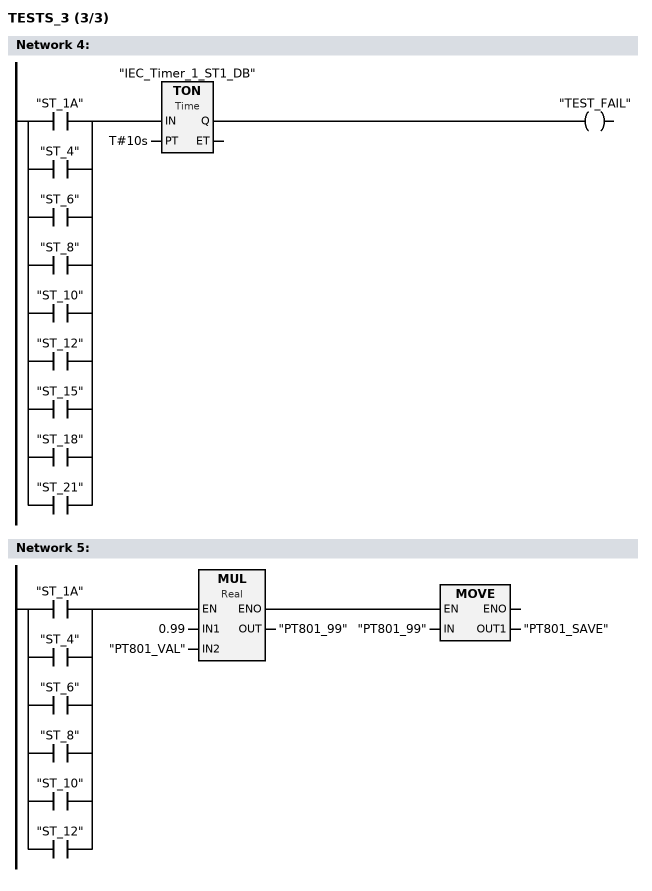
   "IEC_Timer_1_ST1_DB".TON(IN := "ST_1A" OR "ST_4" OR "ST_6" OR "ST_8" OR "ST_10" OR "ST_12" OR "ST_15" OR "ST_18" OR "ST_21",
                           PT := T#10s);
   "TEST_FAIL" := "IEC_Timer_1_ST1_DB".Q;
END_REGION

REGION Network 5
   RUNG wire#powerrail
      Contact( "ST_1A" )
      wire#w1
      { S7_Templates := "SrcType := Real" } Mul(in1 := 0.99, in2 := "PT801_VAL", out => "PT801_99")
      { S7_GenerateENO := "TRUE" } Move(in := "PT801_99", out1 => "PT801_SAVE")
   END_RUNG
   RUNG wire#powerrail
      Contact( "ST_4" )
   END_RUNG wire#w1
   RUNG wire#powerrail
      Contact( "ST_6" )
   END_RUNG wire#w1
   RUNG wire#powerrail
      Contact( "ST_8" )
   END_RUNG wire#w1
   RUNG wire#powerrail
      Contact( "ST_10" )
   END_RUNG wire#w1
   RUNG wire#powerrail
      Contact( "ST_12" )
   END_RUNG wire#w1
   // the same network as SCL:
   IF "ST_1A" OR "ST_4" OR "ST_6" OR "ST_8" OR "ST_10" OR "ST_12" THEN
       "PT801_99" := 0.99 * "PT801_VAL";
       "PT801_SAVE" := "PT801_99";
   END_IF;
END_REGION
END_FUNCTION

FUNCTION "TESTS_2" : Void   // FC18, LAD
{ S7_Optimized_Access := 'FALSE' }
VERSION : 0.1
// Test_MFC401
   VAR_TEMP   // added for the SCL form of the ladder/FBD networks
      _w1 : Bool;
      _w2 : Bool;
   END_VAR
BEGIN

REGION Network 1
   // ALARM Settings
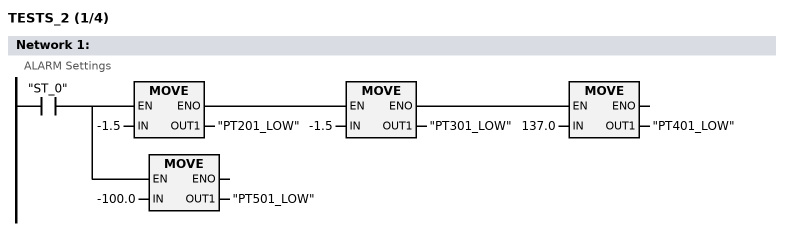
   RUNG wire#powerrail
      Contact( "ST_0" )
      wire#w1
      { S7_GenerateENO := "TRUE" } Move(in := -1.5, out1 => "PT201_LOW")
      { S7_GenerateENO := "TRUE" } Move(in := -1.5, out1 => "PT301_LOW")
      { S7_GenerateENO := "TRUE" } Move(in := 137.0, out1 => "PT401_LOW")
   END_RUNG
   RUNG wire#w1
      { S7_GenerateENO := "TRUE" } Move(in := -100.0, out1 => "PT501_LOW")
   END_RUNG
   // the same network as SCL:
   // ENO of a box is taken as its EN; it also drops when the box reports an error
   IF "ST_0" THEN
       "PT201_LOW" := -1.5;
       "PT301_LOW" := -1.5;
       "PT401_LOW" := 137.0;
       "PT501_LOW" := -100.0;
   END_IF;
END_REGION

REGION Network 2: Pneumatic Tests
   // Test Pneumatic System (Test #1-#6)
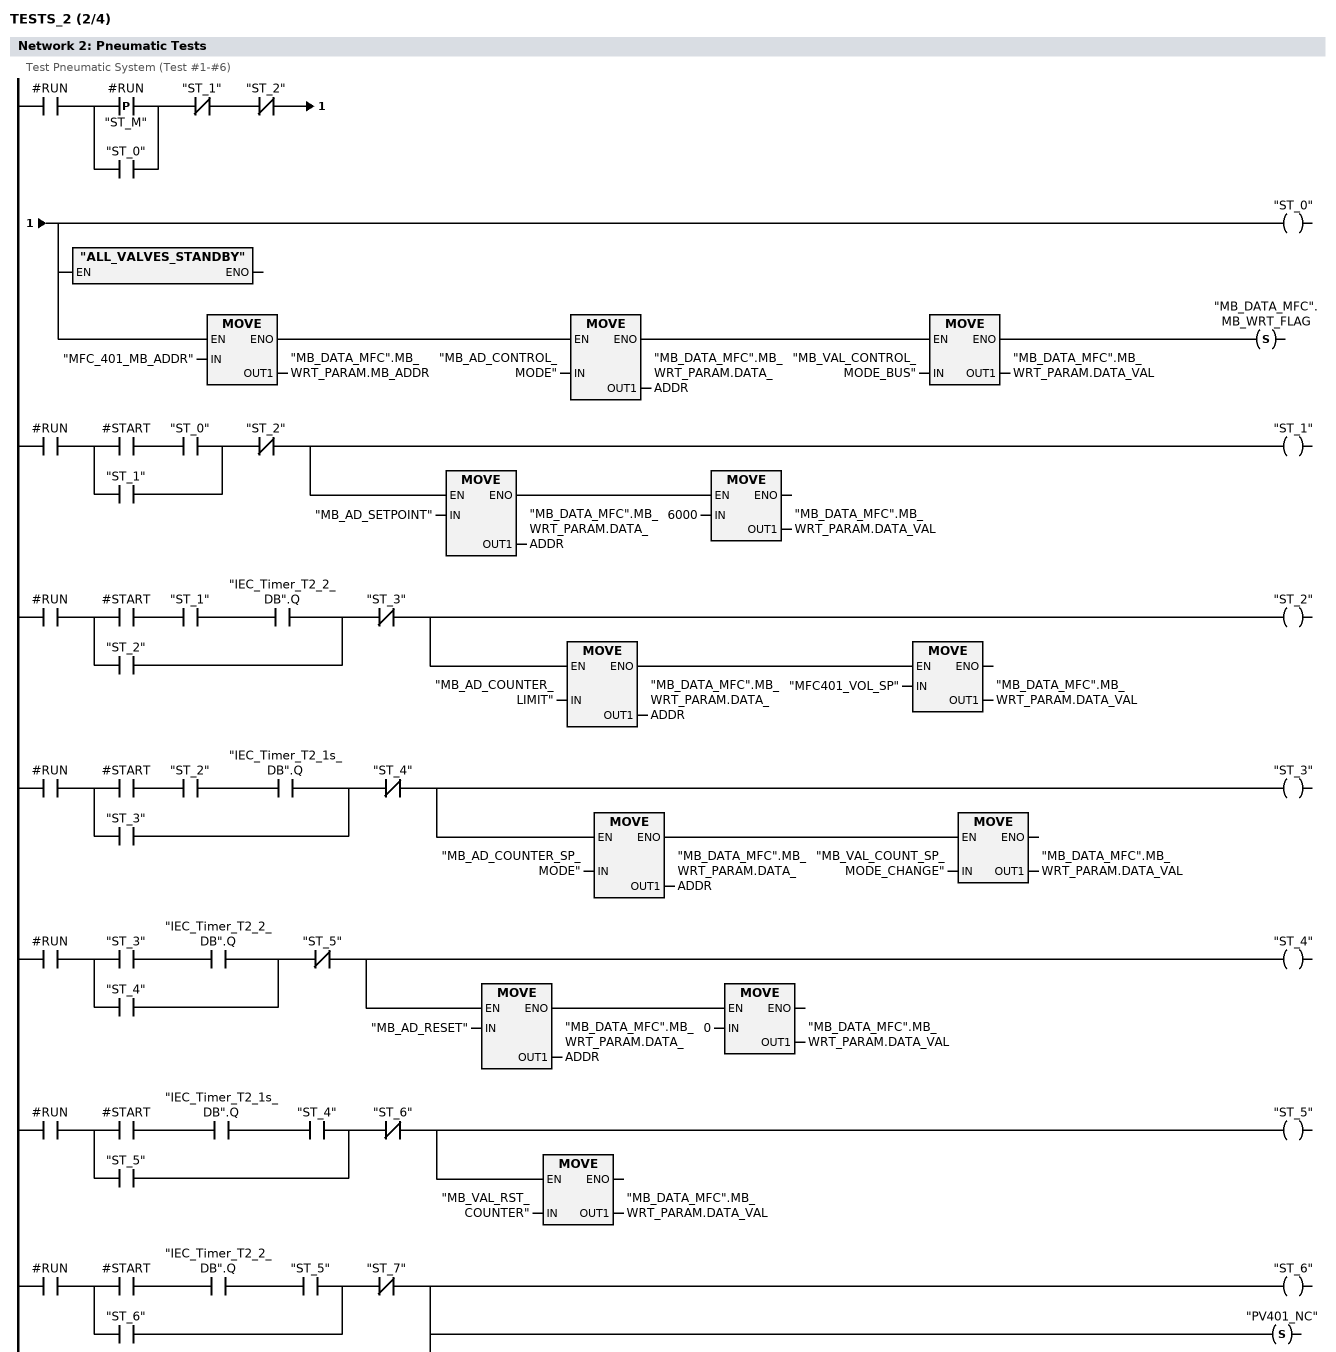
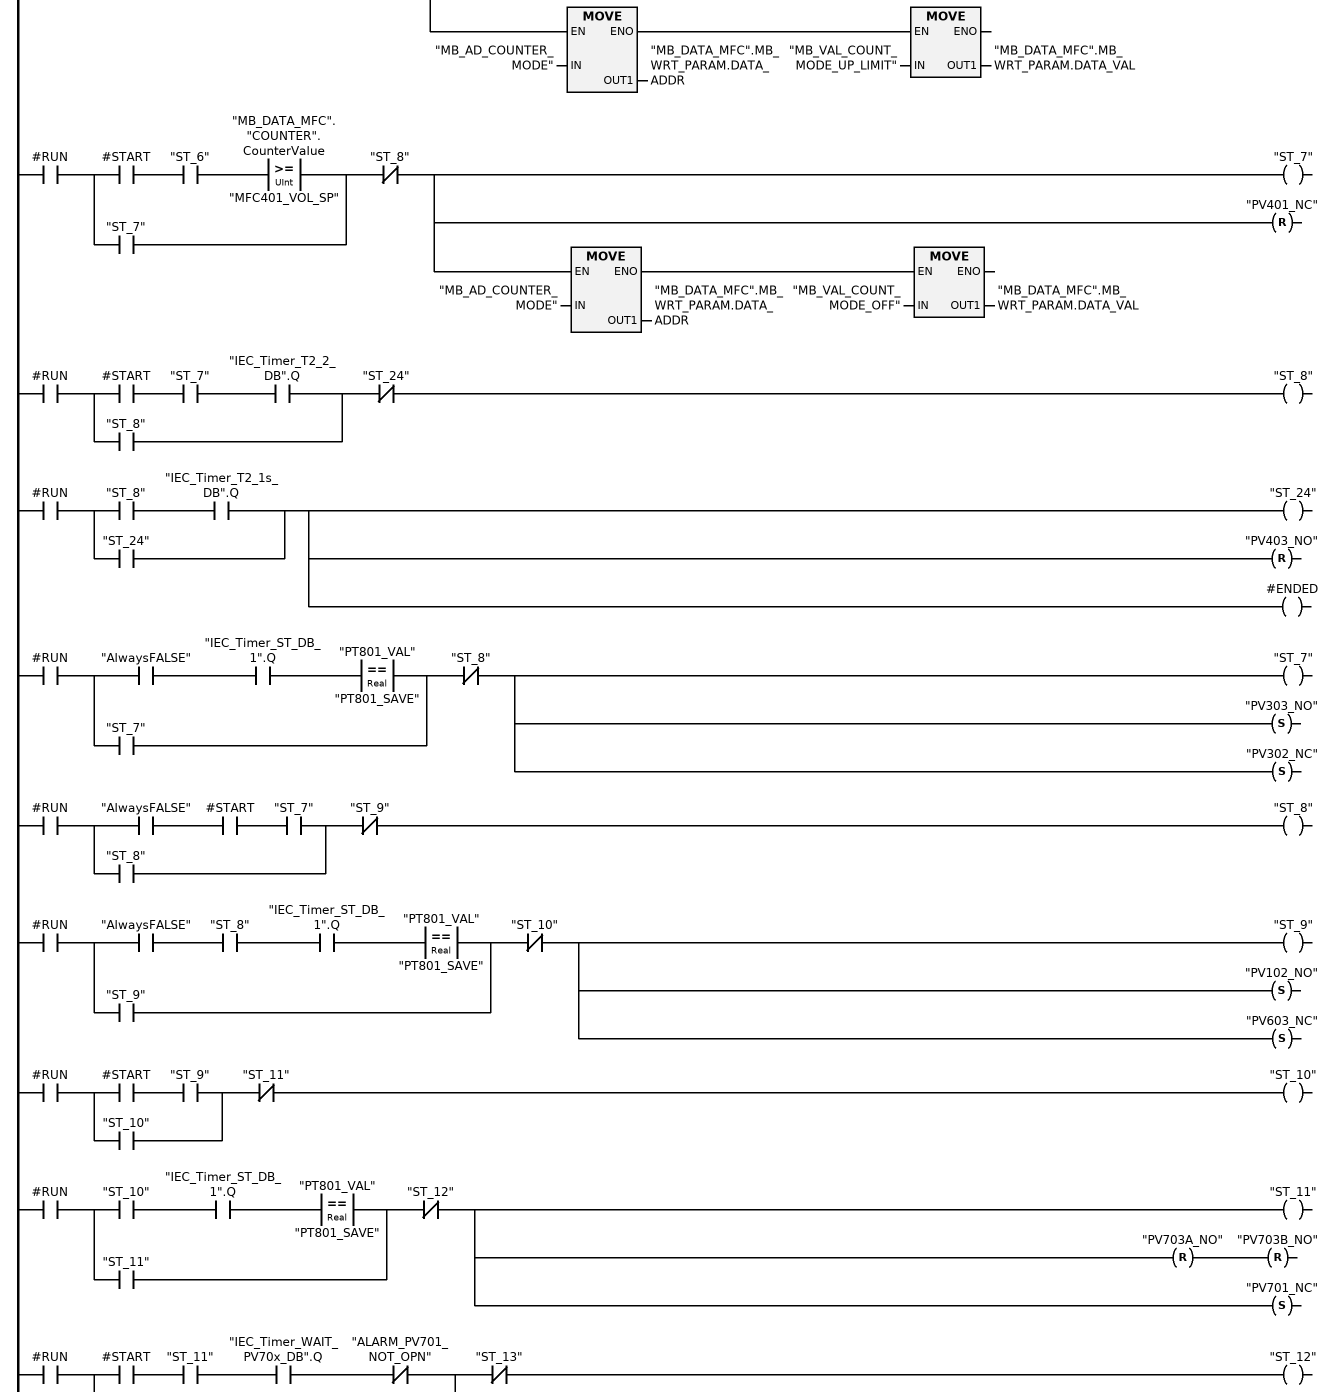
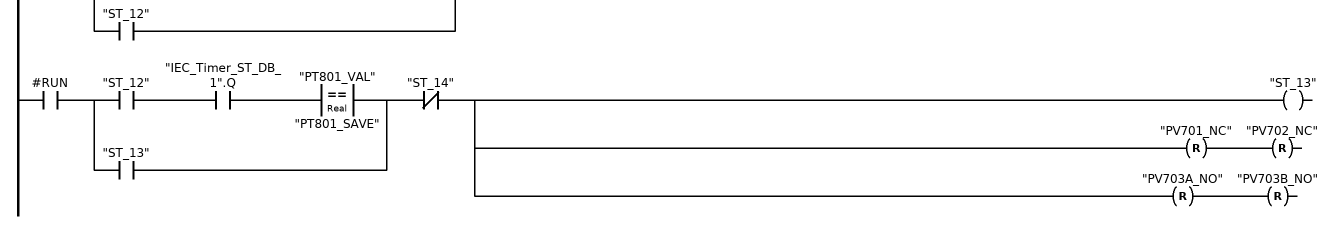
   RUNG wire#powerrail
      Contact( #RUN )
      wire#w1
      P_Contact(operand := #RUN, bit := "ST_M")
      wire#w2
      I_Contact( "ST_1" )
      I_Contact( "ST_2" )
      wire#w3
      Coil( "ST_0" )
   END_RUNG
   RUNG wire#w1
      Contact( "ST_0" )
   END_RUNG wire#w2
   RUNG wire#w3
      "ALL_VALVES_STANDBY"()
   END_RUNG
   RUNG wire#w3
      Move(in := "MFC_401_MB_ADDR", out1 => "MB_DATA_MFC".MB_WRT_PARAM.MB_ADDR)
      Move(in := "MB_AD_CONTROL_MODE", out1 => "MB_DATA_MFC".MB_WRT_PARAM.DATA_ADDR)
      Move(in := "MB_VAL_CONTROL_MODE_BUS", out1 => "MB_DATA_MFC".MB_WRT_PARAM.DATA_VAL)
      S_Coil( "MB_DATA_MFC".MB_WRT_FLAG )
   END_RUNG
   RUNG wire#powerrail
      Contact( #RUN )
      wire#w4
      Contact( #START )
      Contact( "ST_0" )
      wire#w5
      I_Contact( "ST_2" )
      wire#w6
      Coil( "ST_1" )
   END_RUNG
   RUNG wire#w4
      Contact( "ST_1" )
   END_RUNG wire#w5
   RUNG wire#w6
      Move(in := "MB_AD_SETPOINT", out1 => "MB_DATA_MFC".MB_WRT_PARAM.DATA_ADDR)
      Move(in := 6000, out1 => "MB_DATA_MFC".MB_WRT_PARAM.DATA_VAL)
   END_RUNG
   RUNG wire#powerrail
      Contact( #RUN )
      wire#w7
      Contact( #START )
      Contact( "ST_1" )
      Contact( "IEC_Timer_T2_2_DB".Q )
      wire#w8
      I_Contact( "ST_3" )
      wire#w9
      Coil( "ST_2" )
   END_RUNG
   RUNG wire#w7
      Contact( "ST_2" )
   END_RUNG wire#w8
   RUNG wire#w9
      Move(in := "MB_AD_COUNTER_LIMIT", out1 => "MB_DATA_MFC".MB_WRT_PARAM.DATA_ADDR)
      Move(in := "MFC401_VOL_SP", out1 => "MB_DATA_MFC".MB_WRT_PARAM.DATA_VAL)
   END_RUNG
   RUNG wire#powerrail
      Contact( #RUN )
      wire#w10
      Contact( #START )
      Contact( "ST_2" )
      Contact( "IEC_Timer_T2_1s_DB".Q )
      wire#w11
      I_Contact( "ST_4" )
      wire#w12
      Coil( "ST_3" )
   END_RUNG
   RUNG wire#w10
      Contact( "ST_3" )
   END_RUNG wire#w11
   RUNG wire#w12
      Move(in := "MB_AD_COUNTER_SP_MODE", out1 => "MB_DATA_MFC".MB_WRT_PARAM.DATA_ADDR)
      Move(in := "MB_VAL_COUNT_SP_MODE_CHANGE", out1 => "MB_DATA_MFC".MB_WRT_PARAM.DATA_VAL)
   END_RUNG
   RUNG wire#powerrail
      Contact( #RUN )
      wire#w13
      Contact( "ST_3" )
      Contact( "IEC_Timer_T2_2_DB".Q )
      wire#w14
      I_Contact( "ST_5" )
      wire#w15
      Coil( "ST_4" )
   END_RUNG
   RUNG wire#w13
      Contact( "ST_4" )
   END_RUNG wire#w14
   RUNG wire#w15
      Move(in := "MB_AD_RESET", out1 => "MB_DATA_MFC".MB_WRT_PARAM.DATA_ADDR)
      Move(in := 0, out1 => "MB_DATA_MFC".MB_WRT_PARAM.DATA_VAL)
   END_RUNG
   RUNG wire#powerrail
      Contact( #RUN )
      wire#w16
      Contact( #START )
      Contact( "IEC_Timer_T2_1s_DB".Q )
      Contact( "ST_4" )
      wire#w17
      I_Contact( "ST_6" )
      wire#w18
      Coil( "ST_5" )
   END_RUNG
   RUNG wire#w16
      Contact( "ST_5" )
   END_RUNG wire#w17
   RUNG wire#w18
      Move(in := "MB_VAL_RST_COUNTER", out1 => "MB_DATA_MFC".MB_WRT_PARAM.DATA_VAL)
   END_RUNG
   RUNG wire#powerrail
      Contact( #RUN )
      wire#w19
      Contact( #START )
      Contact( "IEC_Timer_T2_2_DB".Q )
      Contact( "ST_5" )
      wire#w20
      I_Contact( "ST_7" )
      wire#w21
      Coil( "ST_6" )
   END_RUNG
   RUNG wire#w19
      Contact( "ST_6" )
   END_RUNG wire#w20
   RUNG wire#w21
      S_Coil( "PV401_NC" )
   END_RUNG
   RUNG wire#w21
      Move(in := "MB_AD_COUNTER_MODE", out1 => "MB_DATA_MFC".MB_WRT_PARAM.DATA_ADDR)
      Move(in := "MB_VAL_COUNT_MODE_UP_LIMIT", out1 => "MB_DATA_MFC".MB_WRT_PARAM.DATA_VAL)
   END_RUNG
   RUNG wire#powerrail
      Contact( #RUN )
      wire#w22
      Contact( #START )
      Contact( "ST_6" )
      { S7_Templates := "SrcType := UInt" } GE_Contact(in1 := "MB_DATA_MFC"."COUNTER".CounterValue, in2 := "MFC401_VOL_SP")
      wire#w23
      I_Contact( "ST_8" )
      wire#w24
      Coil( "ST_7" )
   END_RUNG
   RUNG wire#w22
      Contact( "ST_7" )
   END_RUNG wire#w23
   RUNG wire#w24
      R_Coil( "PV401_NC" )
   END_RUNG
   RUNG wire#w24
      Move(in := "MB_AD_COUNTER_MODE", out1 => "MB_DATA_MFC".MB_WRT_PARAM.DATA_ADDR)
      Move(in := "MB_VAL_COUNT_MODE_OFF", out1 => "MB_DATA_MFC".MB_WRT_PARAM.DATA_VAL)
   END_RUNG
   RUNG wire#powerrail
      Contact( #RUN )
      wire#w25
      Contact( #START )
      Contact( "ST_7" )
      Contact( "IEC_Timer_T2_2_DB".Q )
      wire#w26
      I_Contact( "ST_24" )
      Coil( "ST_8" )
   END_RUNG
   RUNG wire#w25
      Contact( "ST_8" )
   END_RUNG wire#w26
   RUNG wire#powerrail
      Contact( #RUN )
      wire#w27
      Contact( "ST_8" )
      Contact( "IEC_Timer_T2_1s_DB".Q )
      wire#w28
      Coil( "ST_24" )
   END_RUNG
   RUNG wire#w27
      Contact( "ST_24" )
   END_RUNG wire#w28
   RUNG wire#w28
      R_Coil( "PV403_NO" )
   END_RUNG
   RUNG wire#w28
      Coil( #ENDED )
   END_RUNG
   RUNG wire#powerrail
      Contact( #RUN )
      wire#w29
      Contact( "AlwaysFALSE" )
      Contact( "IEC_Timer_ST_DB_1".Q )
      { S7_Templates := "SrcType := Real" } EQ_Contact(in1 := "PT801_VAL", in2 := "PT801_SAVE")
      wire#w30
      I_Contact( "ST_8" )
      wire#w31
      Coil( "ST_7" )
   END_RUNG
   RUNG wire#w29
      Contact( "ST_7" )
   END_RUNG wire#w30
   RUNG wire#w31
      S_Coil( "PV303_NO" )
   END_RUNG
   RUNG wire#w31
      S_Coil( "PV302_NC" )
   END_RUNG
   RUNG wire#powerrail
      Contact( #RUN )
      wire#w32
      Contact( "AlwaysFALSE" )
      Contact( #START )
      Contact( "ST_7" )
      wire#w33
      I_Contact( "ST_9" )
      Coil( "ST_8" )
   END_RUNG
   RUNG wire#w32
      Contact( "ST_8" )
   END_RUNG wire#w33
   RUNG wire#powerrail
      Contact( #RUN )
      wire#w34
      Contact( "AlwaysFALSE" )
      Contact( "ST_8" )
      Contact( "IEC_Timer_ST_DB_1".Q )
      { S7_Templates := "SrcType := Real" } EQ_Contact(in1 := "PT801_VAL", in2 := "PT801_SAVE")
      wire#w35
      I_Contact( "ST_10" )
      wire#w36
      Coil( "ST_9" )
   END_RUNG
   RUNG wire#w34
      Contact( "ST_9" )
   END_RUNG wire#w35
   RUNG wire#w36
      S_Coil( "PV102_NO" )
   END_RUNG
   RUNG wire#w36
      S_Coil( "PV603_NC" )
   END_RUNG
   RUNG wire#powerrail
      Contact( #RUN )
      wire#w37
      Contact( #START )
      Contact( "ST_9" )
      wire#w38
      I_Contact( "ST_11" )
      Coil( "ST_10" )
   END_RUNG
   RUNG wire#w37
      Contact( "ST_10" )
   END_RUNG wire#w38
   RUNG wire#powerrail
      Contact( #RUN )
      wire#w39
      Contact( "ST_10" )
      Contact( "IEC_Timer_ST_DB_1".Q )
      { S7_Templates := "SrcType := Real" } EQ_Contact(in1 := "PT801_VAL", in2 := "PT801_SAVE")
      wire#w40
      I_Contact( "ST_12" )
      wire#w41
      Coil( "ST_11" )
   END_RUNG
   RUNG wire#w39
      Contact( "ST_11" )
   END_RUNG wire#w40
   RUNG wire#w41
      R_Coil( "PV703A_NO" )
      R_Coil( "PV703B_NO" )
   END_RUNG
   RUNG wire#w41
      S_Coil( "PV701_NC" )
   END_RUNG
   RUNG wire#powerrail
      Contact( #RUN )
      wire#w42
      Contact( #START )
      Contact( "ST_11" )
      Contact( "IEC_Timer_WAIT_PV70x_DB".Q )
      I_Contact( "ALARM_PV701_NOT_OPN" )
      wire#w43
      I_Contact( "ST_13" )
      Coil( "ST_12" )
   END_RUNG
   RUNG wire#w42
      Contact( "ST_12" )
   END_RUNG wire#w43
   RUNG wire#powerrail
      Contact( #RUN )
      wire#w44
      Contact( "ST_12" )
      Contact( "IEC_Timer_ST_DB_1".Q )
      { S7_Templates := "SrcType := Real" } EQ_Contact(in1 := "PT801_VAL", in2 := "PT801_SAVE")
      wire#w45
      I_Contact( "ST_14" )
      wire#w46
      Coil( "ST_13" )
   END_RUNG
   RUNG wire#w44
      Contact( "ST_13" )
   END_RUNG wire#w45
   RUNG wire#w46
      R_Coil( "PV701_NC" )
      R_Coil( "PV702_NC" )
   END_RUNG
   RUNG wire#w46
      R_Coil( "PV703A_NO" )
      R_Coil( "PV703B_NO" )
   END_RUNG
   // the same network as SCL:
   #_w1 := #RUN AND #RUN AND NOT "ST_M";   // rising edge of #RUN
   "ST_M" := #RUN;
   "ST_0" := (#_w1 OR (#RUN AND "ST_0")) AND NOT "ST_1" AND NOT "ST_2";
   #_w2 := "ST_0";
   IF #_w2 THEN
       "ALL_VALVES_STANDBY"();
       "MB_DATA_MFC".MB_WRT_PARAM.MB_ADDR := "MFC_401_MB_ADDR";
       "MB_DATA_MFC".MB_WRT_PARAM.DATA_ADDR := "MB_AD_CONTROL_MODE";
       "MB_DATA_MFC".MB_WRT_PARAM.DATA_VAL := "MB_VAL_CONTROL_MODE_BUS";
       "MB_DATA_MFC".MB_WRT_FLAG := TRUE;
   END_IF;
   "ST_1" := #RUN AND ((#START AND "ST_0") OR "ST_1") AND NOT "ST_2";
   IF "ST_1" THEN
       "MB_DATA_MFC".MB_WRT_PARAM.DATA_ADDR := "MB_AD_SETPOINT";
       "MB_DATA_MFC".MB_WRT_PARAM.DATA_VAL := 6000;
   END_IF;
   "ST_2" := #RUN AND ((#START AND "ST_1" AND "IEC_Timer_T2_2_DB".Q) OR "ST_2") AND NOT "ST_3";
   IF "ST_2" THEN
       "MB_DATA_MFC".MB_WRT_PARAM.DATA_ADDR := "MB_AD_COUNTER_LIMIT";
       "MB_DATA_MFC".MB_WRT_PARAM.DATA_VAL := "MFC401_VOL_SP";
   END_IF;
   "ST_3" := #RUN AND ((#START AND "ST_2" AND "IEC_Timer_T2_1s_DB".Q) OR "ST_3") AND NOT "ST_4";
   IF "ST_3" THEN
       "MB_DATA_MFC".MB_WRT_PARAM.DATA_ADDR := "MB_AD_COUNTER_SP_MODE";
       "MB_DATA_MFC".MB_WRT_PARAM.DATA_VAL := "MB_VAL_COUNT_SP_MODE_CHANGE";
   END_IF;
   "ST_4" := #RUN AND (("ST_3" AND "IEC_Timer_T2_2_DB".Q) OR "ST_4") AND NOT "ST_5";
   IF "ST_4" THEN
       "MB_DATA_MFC".MB_WRT_PARAM.DATA_ADDR := "MB_AD_RESET";
       "MB_DATA_MFC".MB_WRT_PARAM.DATA_VAL := 0;
   END_IF;
   "ST_5" := #RUN AND ((#START AND "IEC_Timer_T2_1s_DB".Q AND "ST_4") OR "ST_5") AND NOT "ST_6";
   IF "ST_5" THEN "MB_DATA_MFC".MB_WRT_PARAM.DATA_VAL := "MB_VAL_RST_COUNTER"; END_IF;
   "ST_6" := #RUN AND ((#START AND "IEC_Timer_T2_2_DB".Q AND "ST_5") OR "ST_6") AND NOT "ST_7";
   IF "ST_6" THEN
       "PV401_NC" := TRUE;
       "MB_DATA_MFC".MB_WRT_PARAM.DATA_ADDR := "MB_AD_COUNTER_MODE";
       "MB_DATA_MFC".MB_WRT_PARAM.DATA_VAL := "MB_VAL_COUNT_MODE_UP_LIMIT";
   END_IF;
   "ST_7" := #RUN AND ((#START AND "ST_6" AND ("MB_DATA_MFC"."COUNTER".CounterValue >= "MFC401_VOL_SP")) OR "ST_7") AND NOT "ST_8";
   IF "ST_7" THEN
       "PV401_NC" := FALSE;
       "MB_DATA_MFC".MB_WRT_PARAM.DATA_ADDR := "MB_AD_COUNTER_MODE";
       "MB_DATA_MFC".MB_WRT_PARAM.DATA_VAL := "MB_VAL_COUNT_MODE_OFF";
   END_IF;
   "ST_8" := #RUN AND ((#START AND "ST_7" AND "IEC_Timer_T2_2_DB".Q) OR "ST_8") AND NOT "ST_24";
   "ST_24" := #RUN AND (("ST_8" AND "IEC_Timer_T2_1s_DB".Q) OR "ST_24");
   IF "ST_24" THEN "PV403_NO" := FALSE; END_IF;
   #ENDED := "ST_24";
   "ST_7" := #RUN AND (("AlwaysFALSE" AND "IEC_Timer_ST_DB_1".Q AND ("PT801_VAL" = "PT801_SAVE")) OR "ST_7") AND NOT "ST_8";
   IF "ST_7" THEN
       "PV303_NO" := TRUE;
       "PV302_NC" := TRUE;
   END_IF;
   "ST_8" := #RUN AND (("AlwaysFALSE" AND #START AND "ST_7") OR "ST_8") AND NOT "ST_9";
   "ST_9" := #RUN AND (("AlwaysFALSE" AND "ST_8" AND "IEC_Timer_ST_DB_1".Q AND ("PT801_VAL" = "PT801_SAVE")) OR "ST_9") AND NOT "ST_10";
   IF "ST_9" THEN
       "PV102_NO" := TRUE;
       "PV603_NC" := TRUE;
   END_IF;
   "ST_10" := #RUN AND ((#START AND "ST_9") OR "ST_10") AND NOT "ST_11";
   "ST_11" := #RUN AND (("ST_10" AND "IEC_Timer_ST_DB_1".Q AND ("PT801_VAL" = "PT801_SAVE")) OR "ST_11") AND NOT "ST_12";
   IF "ST_11" THEN
       "PV703A_NO" := FALSE;
       "PV703B_NO" := FALSE;
       "PV701_NC" := TRUE;
   END_IF;
   "ST_12" := #RUN AND ((#START AND "ST_11" AND "IEC_Timer_WAIT_PV70x_DB".Q AND NOT "ALARM_PV701_NOT_OPN") OR "ST_12") AND NOT "ST_13";
   "ST_13" := #RUN AND (("ST_12" AND "IEC_Timer_ST_DB_1".Q AND ("PT801_VAL" = "PT801_SAVE")) OR "ST_13") AND NOT "ST_14";
   IF "ST_13" THEN
       "PV701_NC" := FALSE;
       "PV702_NC" := FALSE;
       "PV703A_NO" := FALSE;
       "PV703B_NO" := FALSE;
   END_IF;
END_REGION

REGION Network 3: Process Tests
   // Tests Process Circuits  (Test #7-#9)
END_REGION

REGION Network 4
   // Timer Wait Test
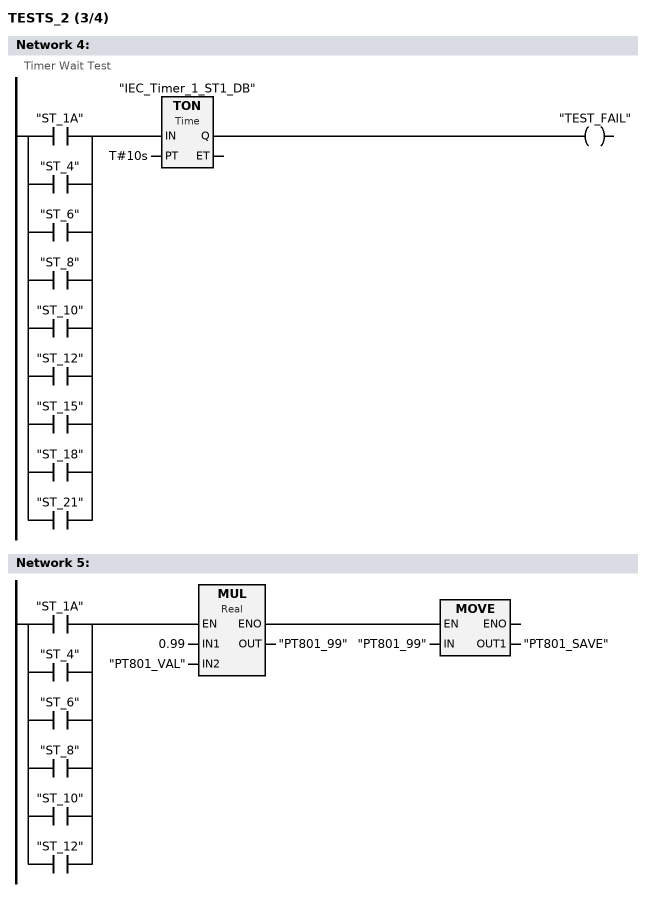
   "IEC_Timer_1_ST1_DB".TON(IN := "ST_1A" OR "ST_4" OR "ST_6" OR "ST_8" OR "ST_10" OR "ST_12" OR "ST_15" OR "ST_18" OR "ST_21",
                           PT := T#10s);
   "TEST_FAIL" := "IEC_Timer_1_ST1_DB".Q;
END_REGION

REGION Network 5
   RUNG wire#powerrail
      Contact( "ST_1A" )
      wire#w1
      { S7_Templates := "SrcType := Real" } Mul(in1 := 0.99, in2 := "PT801_VAL", out => "PT801_99")
      { S7_GenerateENO := "TRUE" } Move(in := "PT801_99", out1 => "PT801_SAVE")
   END_RUNG
   RUNG wire#powerrail
      Contact( "ST_4" )
   END_RUNG wire#w1
   RUNG wire#powerrail
      Contact( "ST_6" )
   END_RUNG wire#w1
   RUNG wire#powerrail
      Contact( "ST_8" )
   END_RUNG wire#w1
   RUNG wire#powerrail
      Contact( "ST_10" )
   END_RUNG wire#w1
   RUNG wire#powerrail
      Contact( "ST_12" )
   END_RUNG wire#w1
   // the same network as SCL:
   IF "ST_1A" OR "ST_4" OR "ST_6" OR "ST_8" OR "ST_10" OR "ST_12" THEN
       "PT801_99" := 0.99 * "PT801_VAL";
       "PT801_SAVE" := "PT801_99";
   END_IF;
END_REGION

REGION Network 6
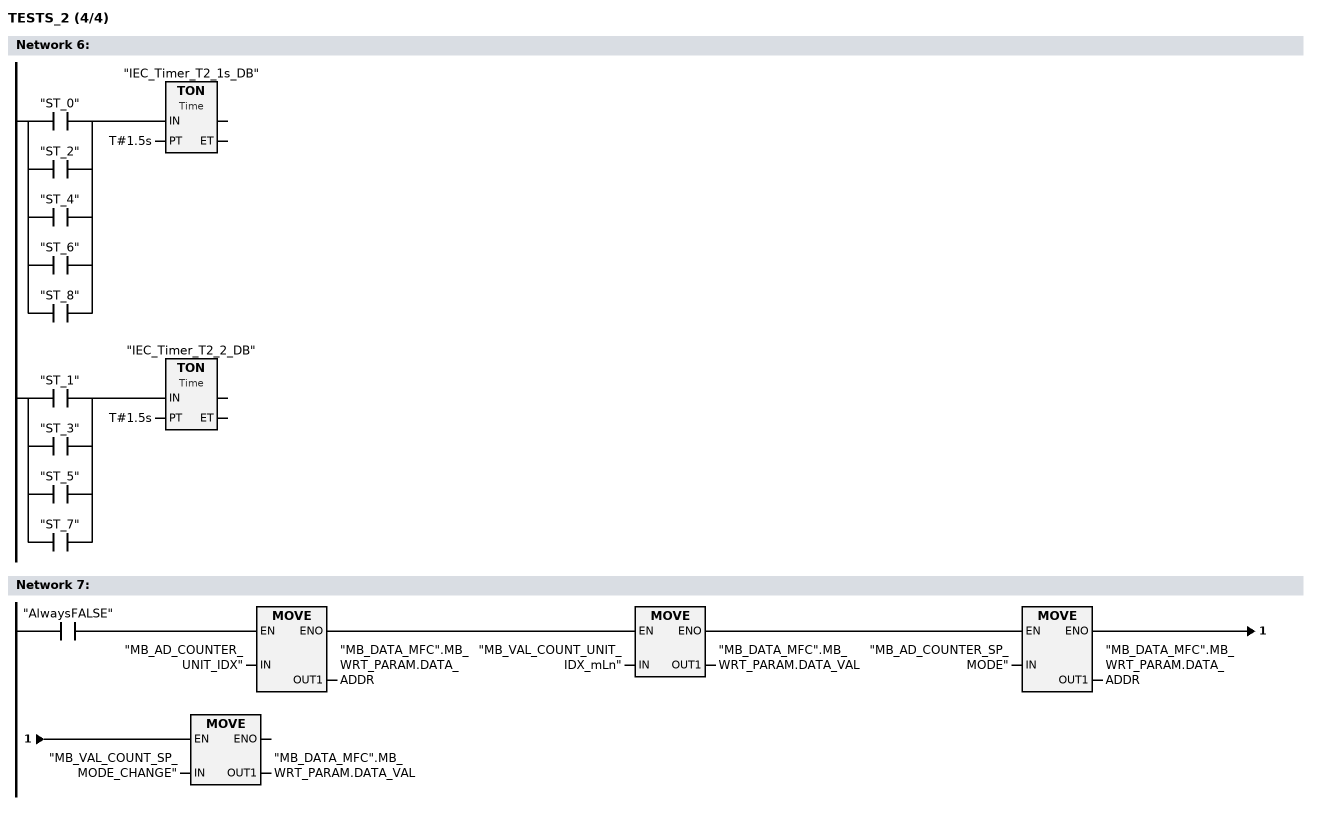
   "IEC_Timer_T2_1s_DB".TON(IN := "ST_0" OR "ST_2" OR "ST_4" OR "ST_6" OR "ST_8", PT := T#1.5s);
   "IEC_Timer_T2_2_DB".TON(IN := "ST_1" OR "ST_3" OR "ST_5" OR "ST_7", PT := T#1.5s);
END_REGION

REGION Network 7
   RUNG wire#powerrail
      Contact( "AlwaysFALSE" )
      Move(in := "MB_AD_COUNTER_UNIT_IDX", out1 => "MB_DATA_MFC".MB_WRT_PARAM.DATA_ADDR)
      Move(in := "MB_VAL_COUNT_UNIT_IDX_mLn", out1 => "MB_DATA_MFC".MB_WRT_PARAM.DATA_VAL)
      Move(in := "MB_AD_COUNTER_SP_MODE", out1 => "MB_DATA_MFC".MB_WRT_PARAM.DATA_ADDR)
      Move(in := "MB_VAL_COUNT_SP_MODE_CHANGE", out1 => "MB_DATA_MFC".MB_WRT_PARAM.DATA_VAL)
   END_RUNG
   // the same network as SCL:
   IF "AlwaysFALSE" THEN
       "MB_DATA_MFC".MB_WRT_PARAM.DATA_ADDR := "MB_AD_COUNTER_UNIT_IDX";
       "MB_DATA_MFC".MB_WRT_PARAM.DATA_VAL := "MB_VAL_COUNT_UNIT_IDX_mLn";
       "MB_DATA_MFC".MB_WRT_PARAM.DATA_ADDR := "MB_AD_COUNTER_SP_MODE";
       "MB_DATA_MFC".MB_WRT_PARAM.DATA_VAL := "MB_VAL_COUNT_SP_MODE_CHANGE";
   END_IF;
END_REGION
END_FUNCTION

FUNCTION "MFC_COUNTER_MODE_SET" : Void   // FC19, LAD
{ S7_Optimized_Access := 'FALSE' }
VERSION : 0.1
   VAR_TEMP   // added for the SCL form of the ladder/FBD networks
      _w1 : Bool;
   END_VAR
BEGIN

REGION Network 1
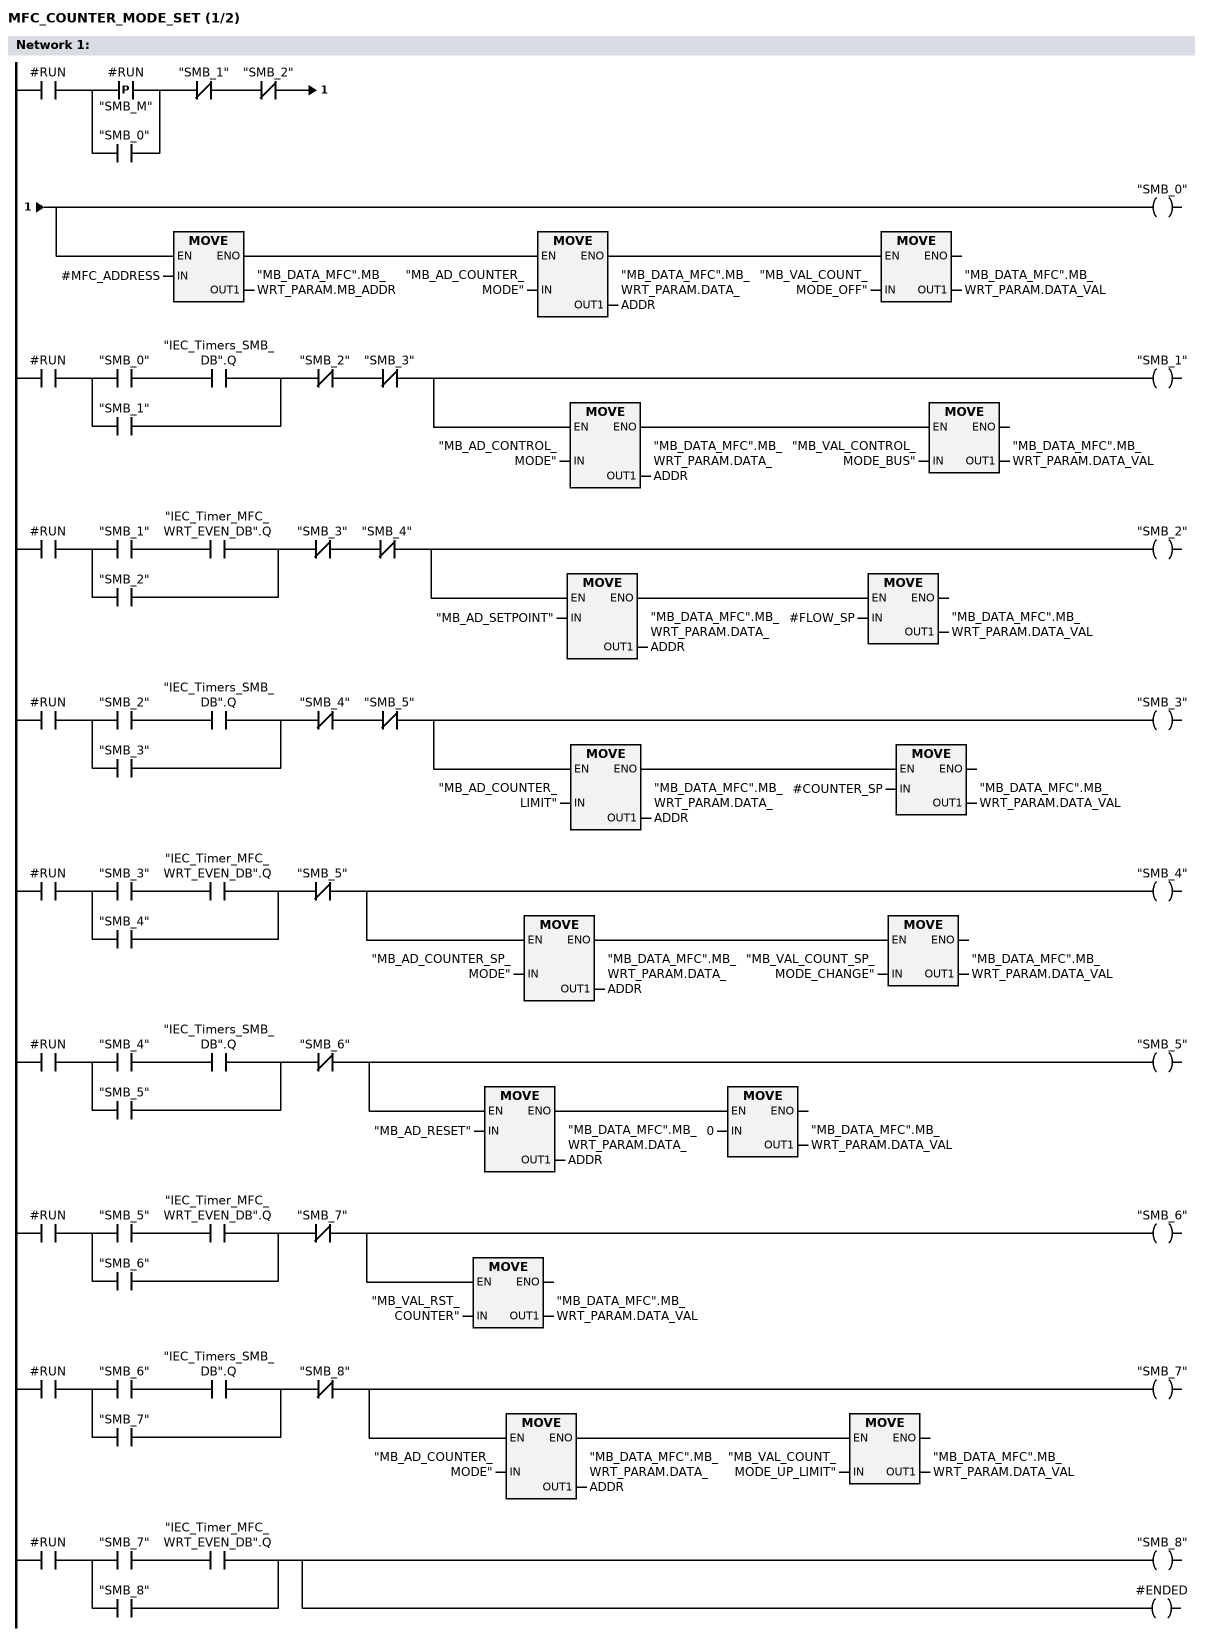
   RUNG wire#powerrail
      Contact( #RUN )
      wire#w1
      P_Contact(operand := #RUN, bit := "SMB_M")
      wire#w2
      I_Contact( "SMB_1" )
      I_Contact( "SMB_2" )
      wire#w3
      Coil( "SMB_0" )
   END_RUNG
   RUNG wire#w1
      Contact( "SMB_0" )
   END_RUNG wire#w2
   RUNG wire#w3
      Move(in := #MFC_ADDRESS, out1 => "MB_DATA_MFC".MB_WRT_PARAM.MB_ADDR)
      Move(in := "MB_AD_COUNTER_MODE", out1 => "MB_DATA_MFC".MB_WRT_PARAM.DATA_ADDR)
      Move(in := "MB_VAL_COUNT_MODE_OFF", out1 => "MB_DATA_MFC".MB_WRT_PARAM.DATA_VAL)
   END_RUNG
   RUNG wire#powerrail
      Contact( #RUN )
      wire#w4
      Contact( "SMB_0" )
      Contact( "IEC_Timers_SMB_DB".Q )
      wire#w5
      I_Contact( "SMB_2" )
      I_Contact( "SMB_3" )
      wire#w6
      Coil( "SMB_1" )
   END_RUNG
   RUNG wire#w4
      Contact( "SMB_1" )
   END_RUNG wire#w5
   RUNG wire#w6
      Move(in := "MB_AD_CONTROL_MODE", out1 => "MB_DATA_MFC".MB_WRT_PARAM.DATA_ADDR)
      Move(in := "MB_VAL_CONTROL_MODE_BUS", out1 => "MB_DATA_MFC".MB_WRT_PARAM.DATA_VAL)
   END_RUNG
   RUNG wire#powerrail
      Contact( #RUN )
      wire#w7
      Contact( "SMB_1" )
      Contact( "IEC_Timer_MFC_WRT_EVEN_DB".Q )
      wire#w8
      I_Contact( "SMB_3" )
      I_Contact( "SMB_4" )
      wire#w9
      Coil( "SMB_2" )
   END_RUNG
   RUNG wire#w7
      Contact( "SMB_2" )
   END_RUNG wire#w8
   RUNG wire#w9
      Move(in := "MB_AD_SETPOINT", out1 => "MB_DATA_MFC".MB_WRT_PARAM.DATA_ADDR)
      Move(in := #FLOW_SP, out1 => "MB_DATA_MFC".MB_WRT_PARAM.DATA_VAL)
   END_RUNG
   RUNG wire#powerrail
      Contact( #RUN )
      wire#w10
      Contact( "SMB_2" )
      Contact( "IEC_Timers_SMB_DB".Q )
      wire#w11
      I_Contact( "SMB_4" )
      I_Contact( "SMB_5" )
      wire#w12
      Coil( "SMB_3" )
   END_RUNG
   RUNG wire#w10
      Contact( "SMB_3" )
   END_RUNG wire#w11
   RUNG wire#w12
      Move(in := "MB_AD_COUNTER_LIMIT", out1 => "MB_DATA_MFC".MB_WRT_PARAM.DATA_ADDR)
      Move(in := #COUNTER_SP, out1 => "MB_DATA_MFC".MB_WRT_PARAM.DATA_VAL)
   END_RUNG
   RUNG wire#powerrail
      Contact( #RUN )
      wire#w13
      Contact( "SMB_3" )
      Contact( "IEC_Timer_MFC_WRT_EVEN_DB".Q )
      wire#w14
      I_Contact( "SMB_5" )
      wire#w15
      Coil( "SMB_4" )
   END_RUNG
   RUNG wire#w13
      Contact( "SMB_4" )
   END_RUNG wire#w14
   RUNG wire#w15
      Move(in := "MB_AD_COUNTER_SP_MODE", out1 => "MB_DATA_MFC".MB_WRT_PARAM.DATA_ADDR)
      Move(in := "MB_VAL_COUNT_SP_MODE_CHANGE", out1 => "MB_DATA_MFC".MB_WRT_PARAM.DATA_VAL)
   END_RUNG
   RUNG wire#powerrail
      Contact( #RUN )
      wire#w16
      Contact( "SMB_4" )
      Contact( "IEC_Timers_SMB_DB".Q )
      wire#w17
      I_Contact( "SMB_6" )
      wire#w18
      Coil( "SMB_5" )
   END_RUNG